(* Logix 5000 project; controller PLC_MCC1300_75F1 vendor 1 type 14 code 166 rev 32.11; software revision 32.04; part 52 of 83 *)
(* tags used below, declared in another part *)
   CONST_rgdDestMask : DINT[32];   // Destination Mask
   CONST_tPlant : UDT_PLANT_CONSTANTS;
   GP_TrackingSearchPlate : GP_TrackingSearchPlate;
   GP_TrackingValidateIndex : GP_TrackingValidateIndex;
   M310_M1_DR_R1 : AXIS_CIP_DRIVE;
   M310_xReqStopPrevConvForPos : BOOL;
   M310Popup : MAC_Popup_ZC[2];
   M310Popup_HMW : MAC_Popup_ZC_HMW[2];
   M310Popup_PlateFreeTimeout : TIMER;
   M310Popup_xDrivePosEnable : BOOL;
   TMP_d : DINT;
   TMP_dDiffPhotocellStartConv0 : DINT;
   TMP_dEndSearch0 : DINT;
   TMP_dEndSearch1 : DINT;
   TMP_dFixedSideOffsetBoth : DINT;
   TMP_dFixedSideOffsetConvoy : DINT;
   TMP_dFixedSideOffsetDW : DINT;
   TMP_dFixedSideOffsetUP : DINT;
   TMP_dHalfConveyorLength : DINT;
   TMP_dHalfPlateLength : DINT;
   TMP_dIndex : DINT;
   TMP_dStartSearch0 : DINT;
   TMP_dStartSearch1 : DINT;
   TMP_xALLForSideLeg : BOOL;
   TMP_xAllLiteToCullet : BOOL;
   TMP_xAtLeastOneForSideLeg : BOOL;
   TMP_xAtLeastOneToCullet : BOOL;
   TMP_xPosHead : BOOL;
   xAlwaysOFF : BOOL;
   xAlwaysON : BOOL;
   xDebugOFF : BOOL;
   Z300_BufferPlate : UDT_LINE_BUFFER_PLATE;
   Z300_Conveyor : UDT_StandConv[29];
   Z300_Conveyor_IN_MOTION : MAC_Conveyor_ZC_IN_MOTION[29];
   Z300_Conveyor_OUT_MOTION : MAC_Conveyor_ZC_OUT_MOTION[29];
   Z300_LineTracking : UDT_LINE_TRACKING;
(* MainProgram, continued *)

ROUTINE M310PopupManagement   (* ladder *)
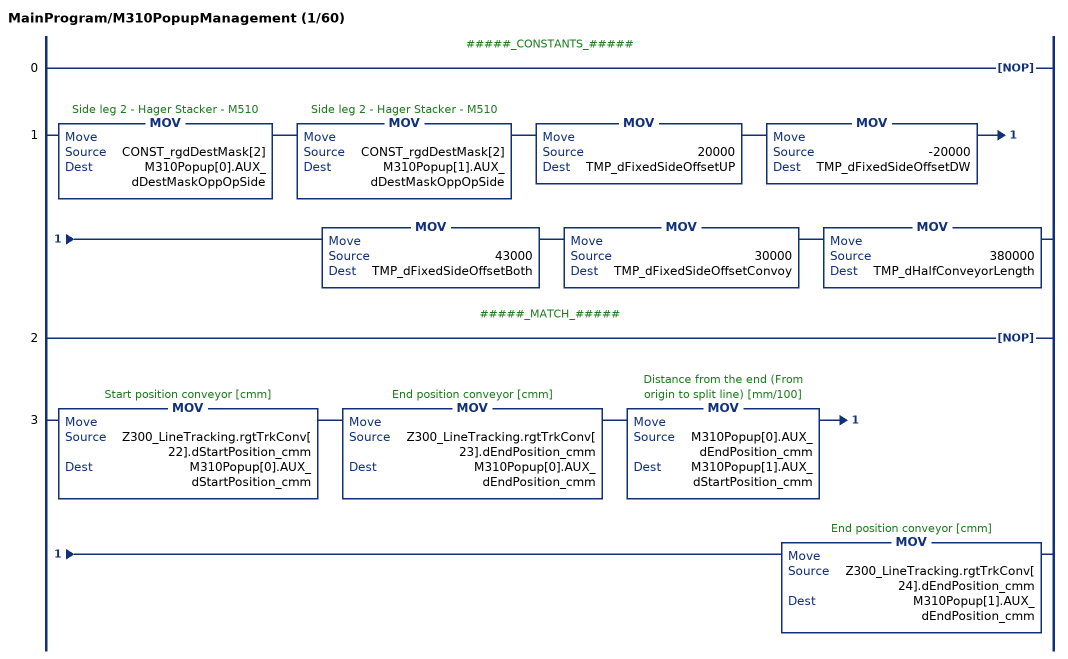
   // #####_CONSTANTS_#####
   0: NOP();
   1: MOV(CONST_rgdDestMask[2],M310Popup[0].AUX_dDestMaskOppOpSide)MOV(CONST_rgdDestMask[2],M310Popup[1].AUX_dDestMaskOppOpSide)MOV(20000,TMP_dFixedSideOffsetUP)MOV(-20000,TMP_dFixedSideOffsetDW)MOV(43000,TMP_dFixedSideOffsetBoth)MOV(30000,TMP_dFixedSideOffsetConvoy)MOV(380000,TMP_dHalfConveyorLength);
   // #####_MATCH_#####
   2: NOP();
   3: MOV(Z300_LineTracking.rgtTrkConv[22].dStartPosition_cmm,M310Popup[0].AUX_dStartPosition_cmm)MOV(Z300_LineTracking.rgtTrkConv[23].dEndPosition_cmm,M310Popup[0].AUX_dEndPosition_cmm)MOV(M310Popup[0].AUX_dEndPosition_cmm,M310Popup[1].AUX_dStartPosition_cmm)MOV(Z300_LineTracking.rgtTrkConv[24].dEndPosition_cmm,M310Popup[1].AUX_dEndPosition_cmm);
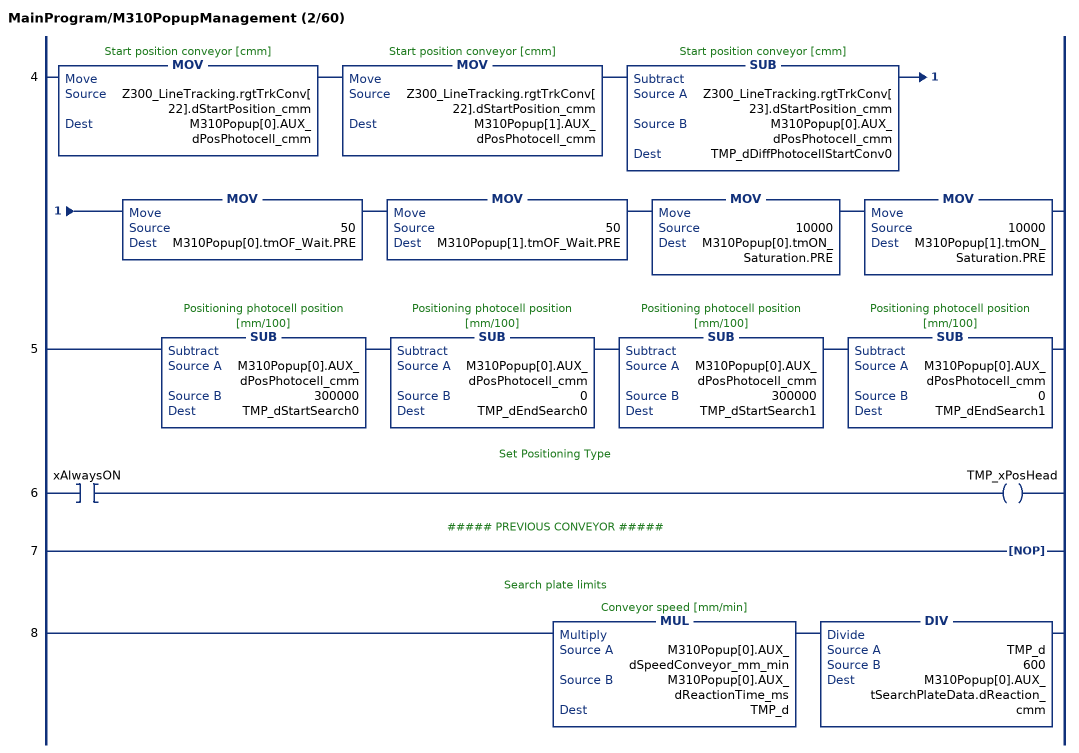
   4: MOV(Z300_LineTracking.rgtTrkConv[22].dStartPosition_cmm,M310Popup[0].AUX_dPosPhotocell_cmm)MOV(Z300_LineTracking.rgtTrkConv[22].dStartPosition_cmm,M310Popup[1].AUX_dPosPhotocell_cmm)SUB(Z300_LineTracking.rgtTrkConv[23].dStartPosition_cmm,M310Popup[0].AUX_dPosPhotocell_cmm,TMP_dDiffPhotocellStartConv0)MOV(50,M310Popup[0].tmOF_Wait.PRE)MOV(50,M310Popup[1].tmOF_Wait.PRE)MOV(10000,M310Popup[0].tmON_Saturation.PRE)MOV(10000,M310Popup[1].tmON_Saturation.PRE);
   5: SUB(M310Popup[0].AUX_dPosPhotocell_cmm,300000,TMP_dStartSearch0)SUB(M310Popup[0].AUX_dPosPhotocell_cmm,0,TMP_dEndSearch0)SUB(M310Popup[0].AUX_dPosPhotocell_cmm,300000,TMP_dStartSearch1)SUB(M310Popup[0].AUX_dPosPhotocell_cmm,0,TMP_dEndSearch1);
   // Set Positioning Type
   6: XIC(xAlwaysON)OTE(TMP_xPosHead);
   // ##### PREVIOUS CONVEYOR #####
   7: NOP();
   // Search plate limits
   8: MUL(M310Popup[0].AUX_dSpeedConveyor_mm_min,M310Popup[0].AUX_dReactionTime_ms,TMP_d)DIV(TMP_d,600,M310Popup[0].AUX_tSearchPlateData.dReaction_cmm);
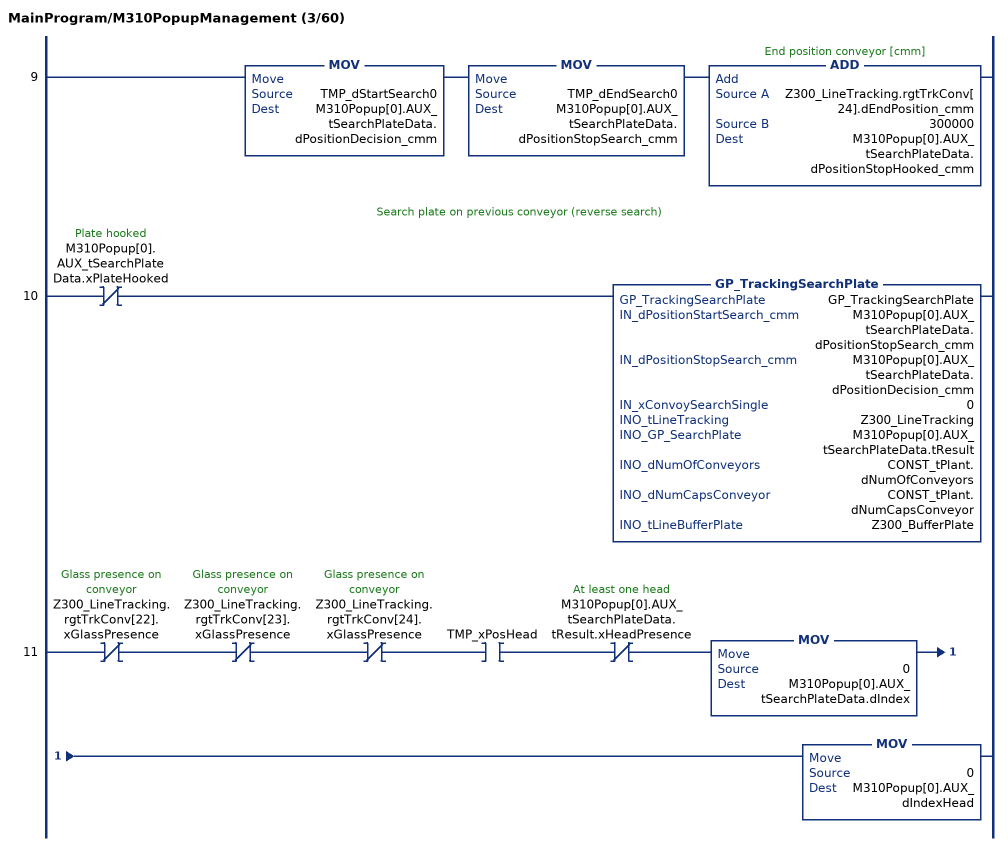
   9: MOV(TMP_dStartSearch0,M310Popup[0].AUX_tSearchPlateData.dPositionDecision_cmm)MOV(TMP_dEndSearch0,M310Popup[0].AUX_tSearchPlateData.dPositionStopSearch_cmm)ADD(Z300_LineTracking.rgtTrkConv[24].dEndPosition_cmm,300000,M310Popup[0].AUX_tSearchPlateData.dPositionStopHooked_cmm);
   // Search plate on previous conveyor (reverse search)
   10: XIO(M310Popup[0].AUX_tSearchPlateData.xPlateHooked)GP_TrackingSearchPlate(GP_TrackingSearchPlate,M310Popup[0].AUX_tSearchPlateData.dPositionStopSearch_cmm,M310Popup[0].AUX_tSearchPlateData.dPositionDecision_cmm,0,Z300_LineTracking,M310Popup[0].AUX_tSearchPlateData.tResult,CONST_tPlant.dNumOfConveyors,CONST_tPlant.dNumCapsConveyor,Z300_BufferPlate);
   11: XIO(Z300_LineTracking.rgtTrkConv[22].xGlassPresence)XIO(Z300_LineTracking.rgtTrkConv[23].xGlassPresence)XIO(Z300_LineTracking.rgtTrkConv[24].xGlassPresence)XIC(TMP_xPosHead)XIO(M310Popup[0].AUX_tSearchPlateData.tResult.xHeadPresence)MOV(0,M310Popup[0].AUX_tSearchPlateData.dIndex)MOV(0,M310Popup[0].AUX_dIndexHead);
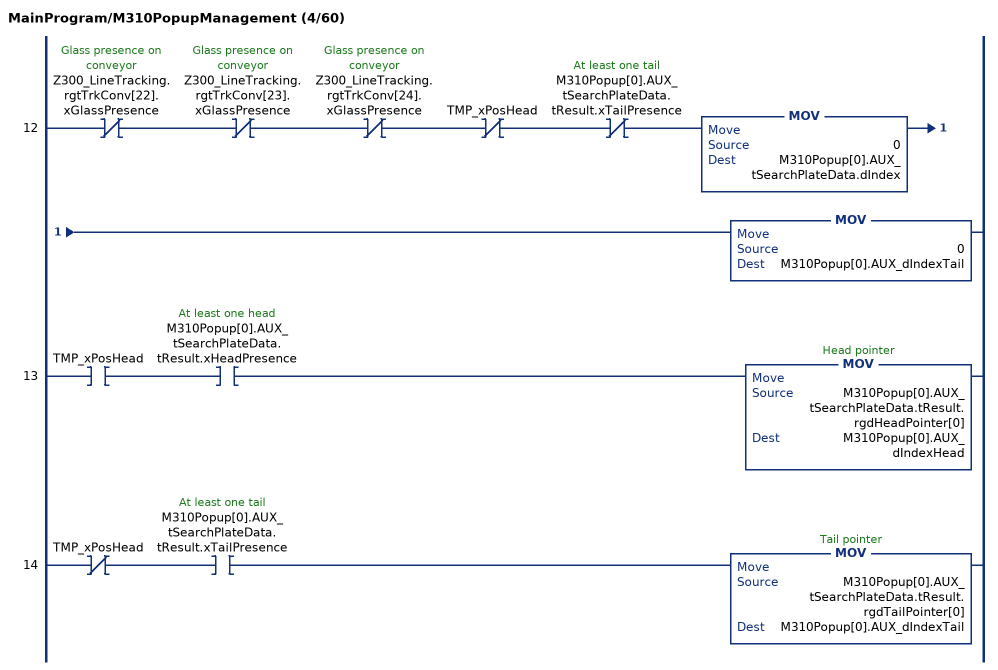
   12: XIO(Z300_LineTracking.rgtTrkConv[22].xGlassPresence)XIO(Z300_LineTracking.rgtTrkConv[23].xGlassPresence)XIO(Z300_LineTracking.rgtTrkConv[24].xGlassPresence)XIO(TMP_xPosHead)XIO(M310Popup[0].AUX_tSearchPlateData.tResult.xTailPresence)MOV(0,M310Popup[0].AUX_tSearchPlateData.dIndex)MOV(0,M310Popup[0].AUX_dIndexTail);
   13: XIC(TMP_xPosHead)XIC(M310Popup[0].AUX_tSearchPlateData.tResult.xHeadPresence)MOV(M310Popup[0].AUX_tSearchPlateData.tResult.rgdHeadPointer[0],M310Popup[0].AUX_dIndexHead);
   14: XIO(TMP_xPosHead)XIC(M310Popup[0].AUX_tSearchPlateData.tResult.xTailPresence)MOV(M310Popup[0].AUX_tSearchPlateData.tResult.rgdTailPointer[0],M310Popup[0].AUX_dIndexTail);
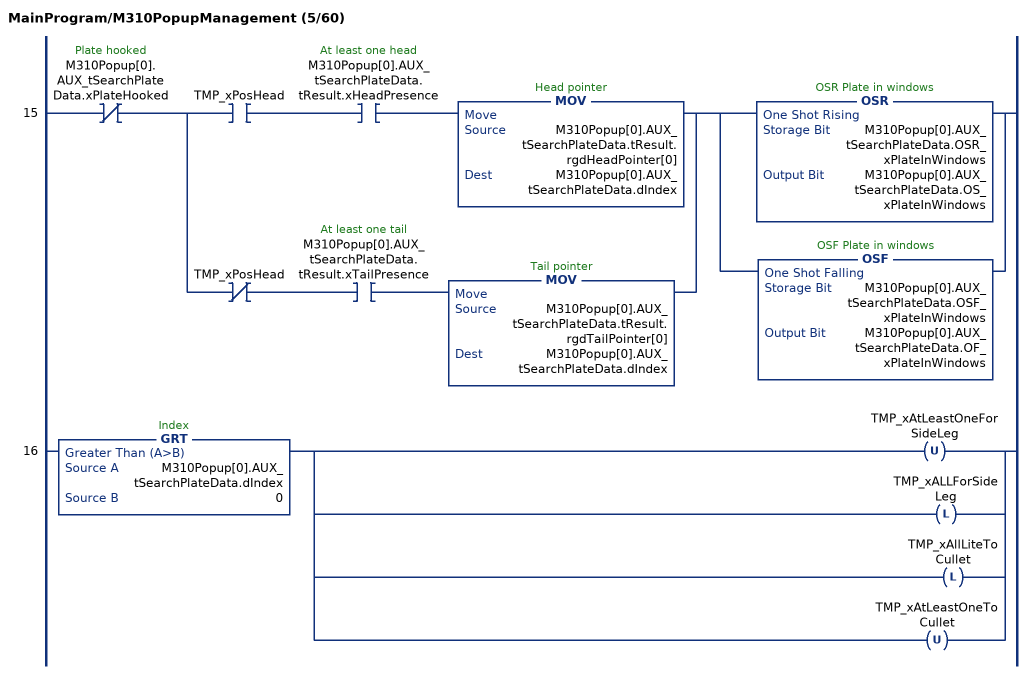
   15: XIO(M310Popup[0].AUX_tSearchPlateData.xPlateHooked)[XIC(TMP_xPosHead) XIC(M310Popup[0].AUX_tSearchPlateData.tResult.xHeadPresence) MOV(M310Popup[0].AUX_tSearchPlateData.tResult.rgdHeadPointer[0],M310Popup[0].AUX_tSearchPlateData.dIndex) ,XIO(TMP_xPosHead) XIC(M310Popup[0].AUX_tSearchPlateData.tResult.xTailPresence) MOV(M310Popup[0].AUX_tSearchPlateData.tResult.rgdTailPointer[0],M310Popup[0].AUX_tSearchPlateData.dIndex) ][OSR(M310Popup[0].AUX_tSearchPlateData.OSR_xPlateInWindows,M310Popup[0].AUX_tSearchPlateData.OS_xPlateInWindows) ,OSF(M310Popup[0].AUX_tSearchPlateData.OSF_xPlateInWindows,M310Popup[0].AUX_tSearchPlateData.OF_xPlateInWindows) ];
   16: GRT(M310Popup[0].AUX_tSearchPlateData.dIndex,0)[OTU(TMP_xAtLeastOneForSideLeg) ,OTL(TMP_xALLForSideLeg) ,OTL(TMP_xAllLiteToCullet) ,OTU(TMP_xAtLeastOneToCullet) ];
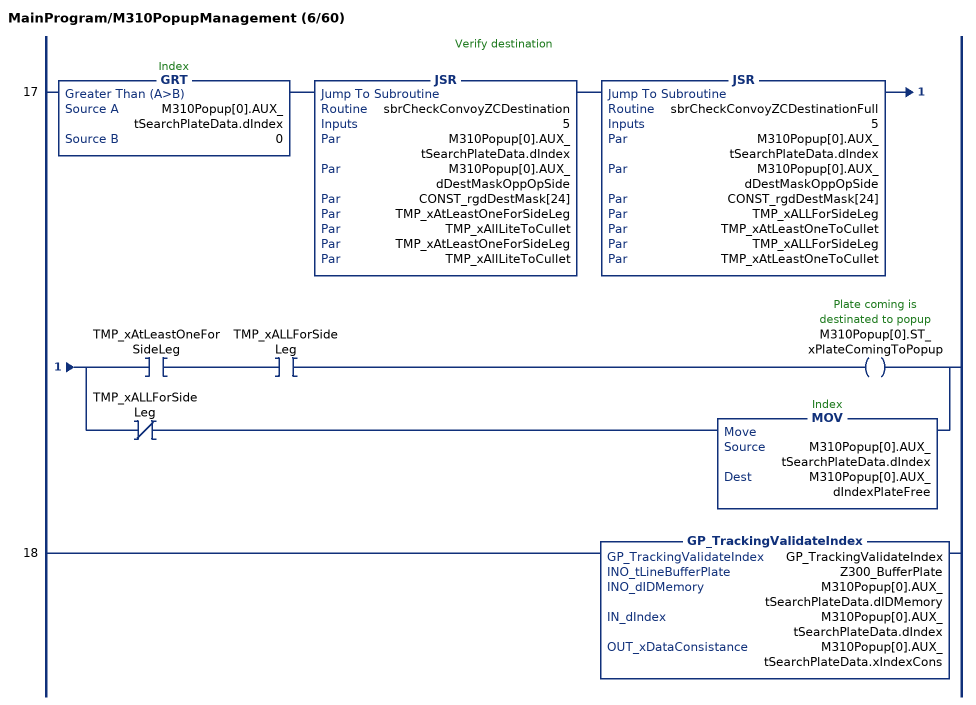
   // Verify destination
   17: GRT(M310Popup[0].AUX_tSearchPlateData.dIndex,0)JSR(sbrCheckConvoyZCDestination,5,M310Popup[0].AUX_tSearchPlateData.dIndex,M310Popup[0].AUX_dDestMaskOppOpSide,CONST_rgdDestMask[24],TMP_xAtLeastOneForSideLeg,TMP_xAllLiteToCullet,TMP_xAtLeastOneForSideLeg,TMP_xAllLiteToCullet)JSR(sbrCheckConvoyZCDestinationFull,5,M310Popup[0].AUX_tSearchPlateData.dIndex,M310Popup[0].AUX_dDestMaskOppOpSide,CONST_rgdDestMask[24],TMP_xALLForSideLeg,TMP_xAtLeastOneToCullet,TMP_xALLForSideLeg,TMP_xAtLeastOneToCullet)[XIC(TMP_xAtLeastOneForSideLeg) XIC(TMP_xALLForSideLeg) OTE(M310Popup[0].ST_xPlateComingToPopup) ,XIO(TMP_xALLForSideLeg) MOV(M310Popup[0].AUX_tSearchPlateData.dIndex,M310Popup[0].AUX_dIndexPlateFree) ];
   18: GP_TrackingValidateIndex(GP_TrackingValidateIndex,Z300_BufferPlate,M310Popup[0].AUX_tSearchPlateData.dIDMemory,M310Popup[0].AUX_tSearchPlateData.dIndex,M310Popup[0].AUX_tSearchPlateData.xIndexCons);
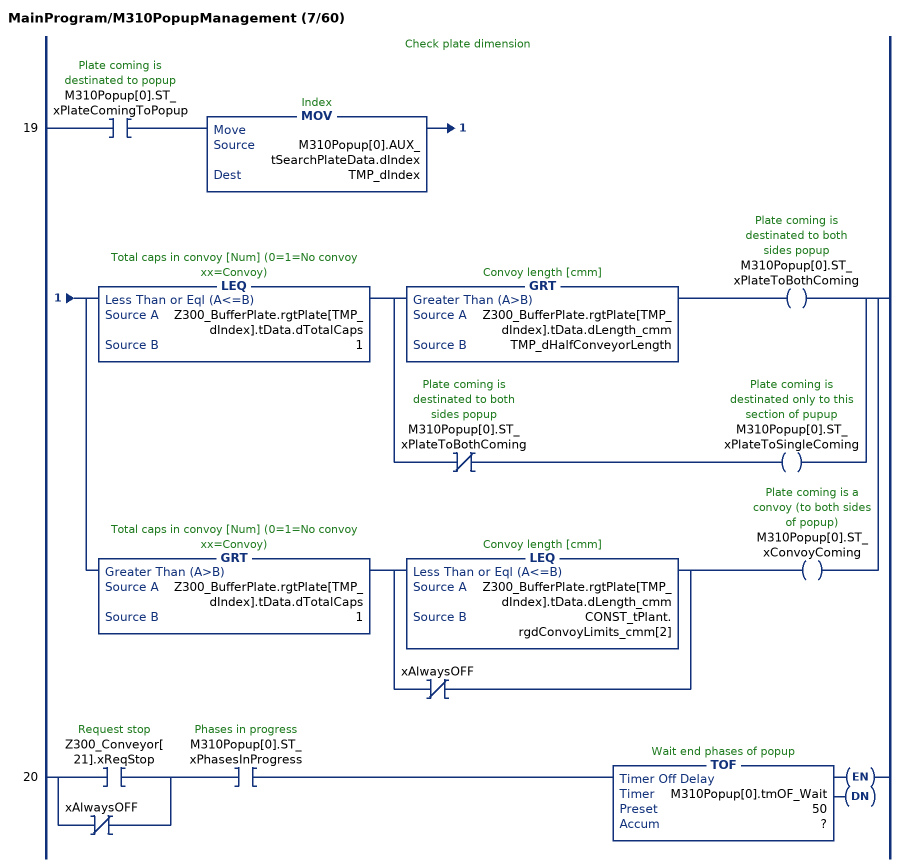
   // Check plate dimension
   19: XIC(M310Popup[0].ST_xPlateComingToPopup)MOV(M310Popup[0].AUX_tSearchPlateData.dIndex,TMP_dIndex)[LEQ(Z300_BufferPlate.rgtPlate[TMP_dIndex].tData.dTotalCaps,1) [GRT(Z300_BufferPlate.rgtPlate[TMP_dIndex].tData.dLength_cmm,TMP_dHalfConveyorLength) OTE(M310Popup[0].ST_xPlateToBothComing) ,XIO(M310Popup[0].ST_xPlateToBothComing) OTE(M310Popup[0].ST_xPlateToSingleComing) ] ,GRT(Z300_BufferPlate.rgtPlate[TMP_dIndex].tData.dTotalCaps,1) [LEQ(Z300_BufferPlate.rgtPlate[TMP_dIndex].tData.dLength_cmm,CONST_tPlant.rgdConvoyLimits_cmm[2]) ,XIO(xAlwaysOFF) ] OTE(M310Popup[0].ST_xConvoyComing) ];
   20: [XIC(Z300_Conveyor[21].xReqStop) ,XIO(xAlwaysOFF) ]XIC(M310Popup[0].ST_xPhasesInProgress)TOF(M310Popup[0].tmOF_Wait,?,?);
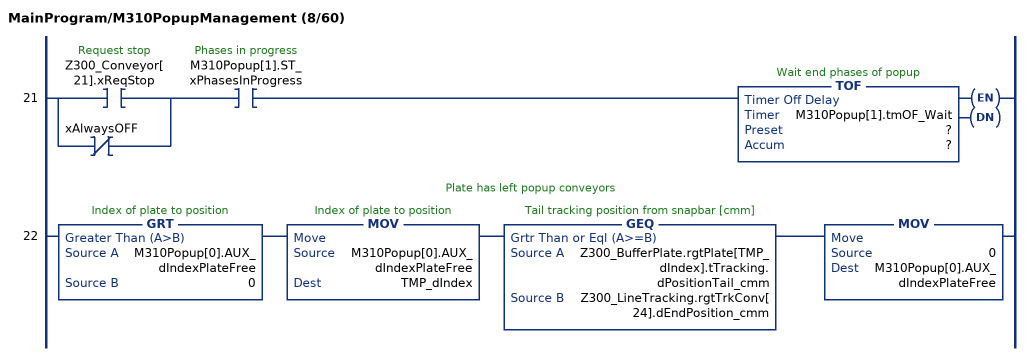
   21: [XIC(Z300_Conveyor[21].xReqStop) ,XIO(xAlwaysOFF) ]XIC(M310Popup[1].ST_xPhasesInProgress)TOF(M310Popup[1].tmOF_Wait,?,?);
   // Plate has left popup conveyors
   22: GRT(M310Popup[0].AUX_dIndexPlateFree,0)MOV(M310Popup[0].AUX_dIndexPlateFree,TMP_dIndex)GEQ(Z300_BufferPlate.rgtPlate[TMP_dIndex].tTracking.dPositionTail_cmm,Z300_LineTracking.rgtTrkConv[24].dEndPosition_cmm)MOV(0,M310Popup[0].AUX_dIndexPlateFree);
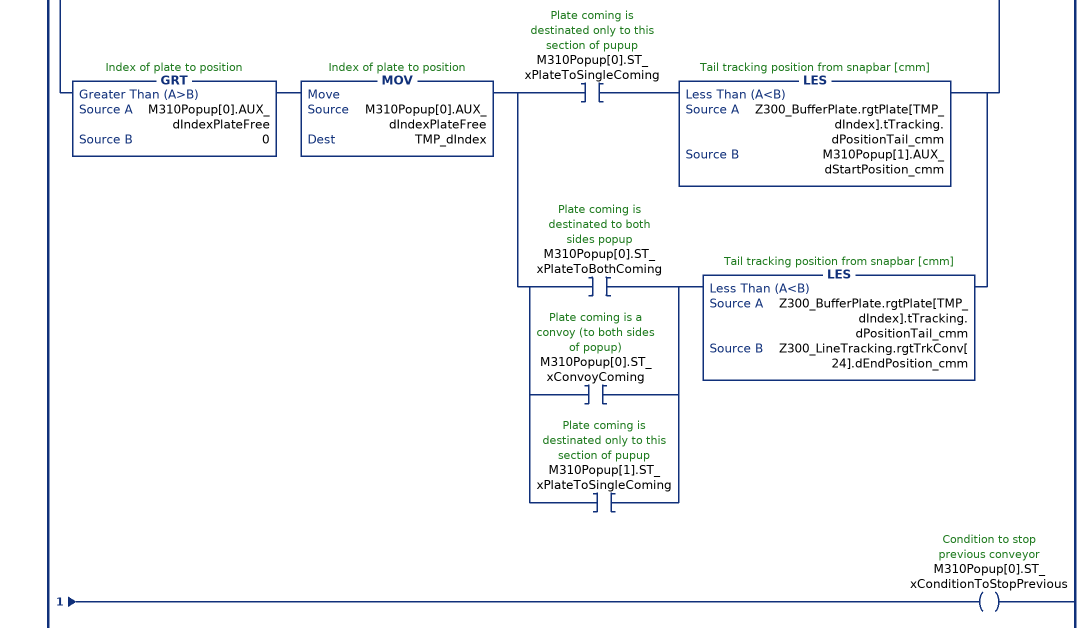
   // Stop previuos conveyor if no condition on pop-up conveyor
   23: [[XIC(M310Popup[0].ST_xPlateToSingleComing) [XIO(M310Popup[0].ST_xInitialConditionForRise) ,XIC(M310Popup[0].ST_xPlatePresentOnPopup) ,XIC(M310Popup[0].ST_xPlatePresence) ,XIC(Z300_LineTracking.rgtTrkConv[22].xGlassPresence) ,XIC(Z300_LineTracking.rgtTrkConv[23].xGlassPresence) ,EQU(M310Popup[0].AUX_dIndexPositioning,0) [XIC(M310Popup[0].ST_xPlateUnderPopup) ,XIC(M310Popup[1].ST_xPlateUnderPopup) ] ] ,XIC(M310Popup[0].ST_xPlateToSingleComing) [XIO(M310Popup[1].ST_xInitialConditionForRise) ,XIC(M310Popup[1].ST_xPlatePresentOnPopup) ,XIC(M310Popup[1].ST_xPlatePresence) ,XIC(Z300_LineTracking.rgtTrkConv[22].xGlassPresence) ,XIC(Z300_LineTracking.rgtTrkConv[23].xGlassPresence) ,XIC(Z300_LineTracking.rgtTrkConv[24].xGlassPresence) ,EQU(M310Popup[0].AUX_dIndexPositioning,0) [XIC(M310Popup[0].ST_xPlateUnderPopup) ,XIC(M310Popup[1].ST_xPlateUnderPopup) ] ] ,[XIC(M310Popup[0].ST_xPlateToBothComing) ,XIC(M310Popup[0].ST_xConvoyComing) ] [XIO(M310Popup[1].ST_xInitialConditionForRise) ,XIC(M310Popup[1].ST_xPlatePresentOnPopup) ,XIC(M310Popup[1].ST_xPlatePresence) ,XIC(Z300_LineTracking.rgtTrkConv[22].xGlassPresence) ,XIC(Z300_LineTracking.rgtTrkConv[23].xGlassPresence) ,XIC(Z300_LineTracking.rgtTrkConv[24].xGlassPresence) ,EQU(M310Popup[0].AUX_dIndexPositioning,0) XIC(M310Popup[1].ST_xPlateUnderPopup) ,XIO(M310Popup[0].ST_xInitialConditionForRise) ,XIC(M310Popup[0].ST_xPlatePresentOnPopup) ,XIC(M310Popup[0].ST_xPlatePresence) ,EQU(M310Popup[0].AUX_dIndexPositioning,0) XIC(M310Popup[0].ST_xPlateUnderPopup) ] ] ,XIO(M310Popup[0].INPUT_xPopupHigh) XIO(M310Popup[0].INPUT_xPopupLow) ,XIO(M310Popup[1].INPUT_xPopupHigh) XIO(M310Popup[1].INPUT_xPopupLow) ,XIC(M310_xReqStopPrevConvForPos) ,XIC(Z300_Conveyor[22].xReqExtStopLoadNewPlate) ,[XIC(M310Popup[0].ST_xPlateInPositionToRise) ,XIC(M310Popup[1].ST_xPlateInPositionToRise) ] ,XIC(Z300_Conveyor[22].ST_xCleaningEnabled) XIO(Z300_Conveyor[21].ST_xCleaningEnabled) ,XIC(M310Popup[0].ST_xPrevConvFreeAfterPos) ,XIC(M310Popup[1].ST_xPrevConvFreeAfterPos) ,[XIO(M310Popup[0].INPUT_xPopupHigh) ,XIO(M310Popup[1].INPUT_xPopupHigh) ] ,GRT(M310Popup[0].AUX_dIndexPositioning,0) [GRT(M310Popup[0].AUX_tSearchPlateData.dIndex,0) NEQ(M310Popup[0].AUX_tSearchPlateData.dIndex,M310Popup[0].AUX_dIndexPositioning) ,GRT(M310Popup[0].AUX_dIndexPlatePositioned,0) NEQ(M310Popup[0].AUX_dIndexPlatePositioned,M310Popup[0].AUX_dIndexPositioning) ] ,GRT(M310Popup[0].AUX_dIndexPlateFree,0) MOV(M310Popup[0].AUX_dIndexPlateFree,TMP_dIndex) [XIC(M310Popup[0].ST_xPlateToSingleComing) LES(Z300_BufferPlate.rgtPlate[TMP_dIndex].tTracking.dPositionTail_cmm,M310Popup[1].AUX_dStartPosition_cmm) ,[XIC(M310Popup[0].ST_xPlateToBothComing) ,XIC(M310Popup[0].ST_xConvoyComing) ,XIC(M310Popup[1].ST_xPlateToSingleComing) ] LES(Z300_BufferPlate.rgtPlate[TMP_dIndex].tTracking.dPositionTail_cmm,Z300_LineTracking.rgtTrkConv[24].dEndPosition_cmm) ] ]OTE(M310Popup[0].ST_xConditionToStopPrevious);
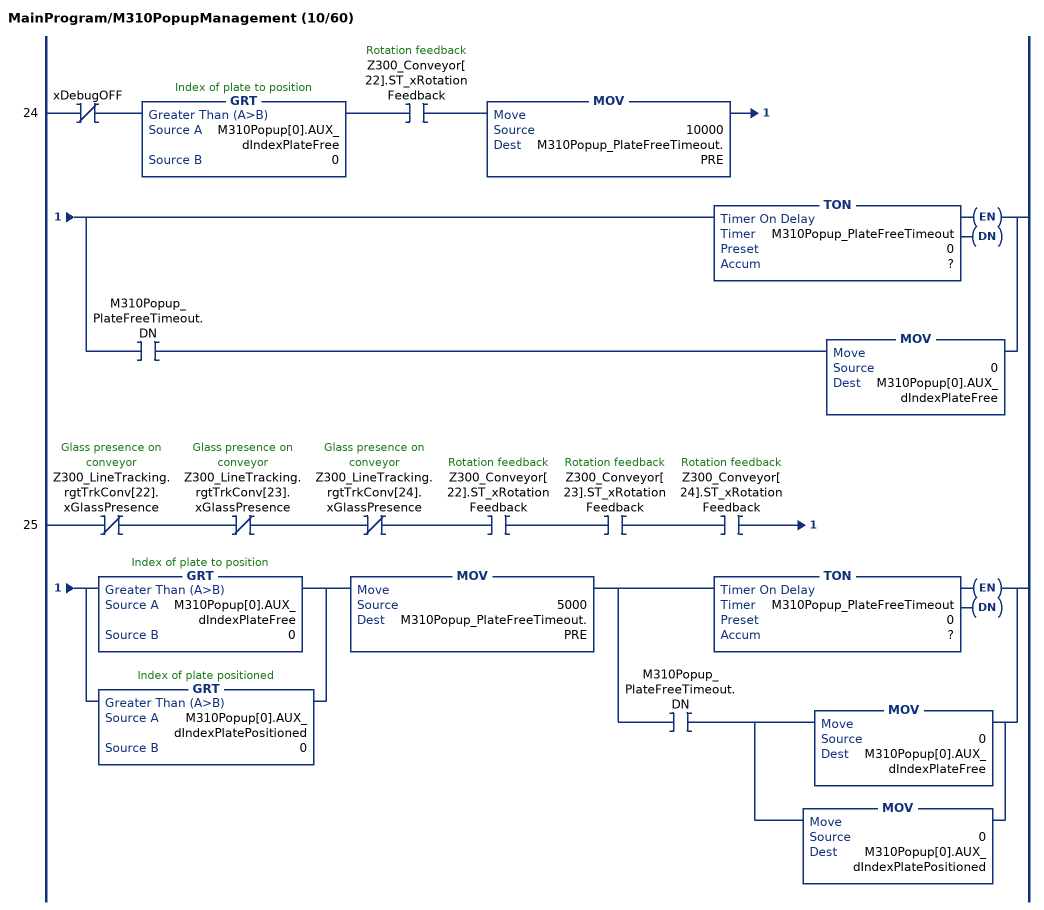
   24: XIO(xDebugOFF)GRT(M310Popup[0].AUX_dIndexPlateFree,0)XIC(Z300_Conveyor[22].ST_xRotationFeedback)MOV(10000,M310Popup_PlateFreeTimeout.PRE)[TON(M310Popup_PlateFreeTimeout,?,?) ,XIC(M310Popup_PlateFreeTimeout.DN) MOV(0,M310Popup[0].AUX_dIndexPlateFree) ];
   25: XIO(Z300_LineTracking.rgtTrkConv[22].xGlassPresence)XIO(Z300_LineTracking.rgtTrkConv[23].xGlassPresence)XIO(Z300_LineTracking.rgtTrkConv[24].xGlassPresence)XIC(Z300_Conveyor[22].ST_xRotationFeedback)XIC(Z300_Conveyor[23].ST_xRotationFeedback)XIC(Z300_Conveyor[24].ST_xRotationFeedback)[GRT(M310Popup[0].AUX_dIndexPlateFree,0) ,GRT(M310Popup[0].AUX_dIndexPlatePositioned,0) ]MOV(5000,M310Popup_PlateFreeTimeout.PRE)[TON(M310Popup_PlateFreeTimeout,?,?) ,XIC(M310Popup_PlateFreeTimeout.DN) [MOV(0,M310Popup[0].AUX_dIndexPlateFree) ,MOV(0,M310Popup[0].AUX_dIndexPlatePositioned) ] ];
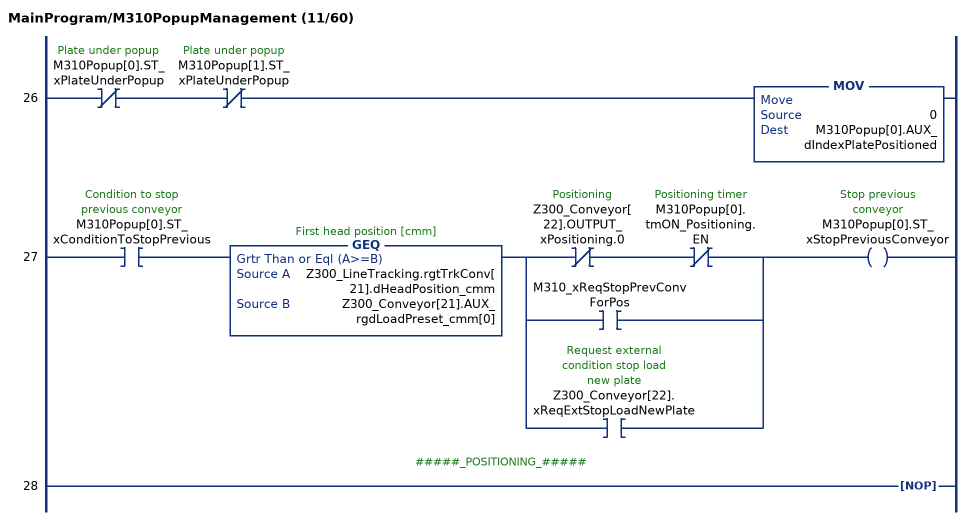
   26: XIO(M310Popup[0].ST_xPlateUnderPopup)XIO(M310Popup[1].ST_xPlateUnderPopup)MOV(0,M310Popup[0].AUX_dIndexPlatePositioned);
   27: XIC(M310Popup[0].ST_xConditionToStopPrevious)GEQ(Z300_LineTracking.rgtTrkConv[21].dHeadPosition_cmm,Z300_Conveyor[21].AUX_rgdLoadPreset_cmm[0])[XIO(Z300_Conveyor[22].OUTPUT_xPositioning.0) XIO(M310Popup[0].tmON_Positioning.EN) ,[XIC(M310_xReqStopPrevConvForPos) ,XIC(Z300_Conveyor[22].xReqExtStopLoadNewPlate) ] ]OTE(M310Popup[0].ST_xStopPreviousConveyor);
   // #####_POSITIONING_#####
   28: NOP();
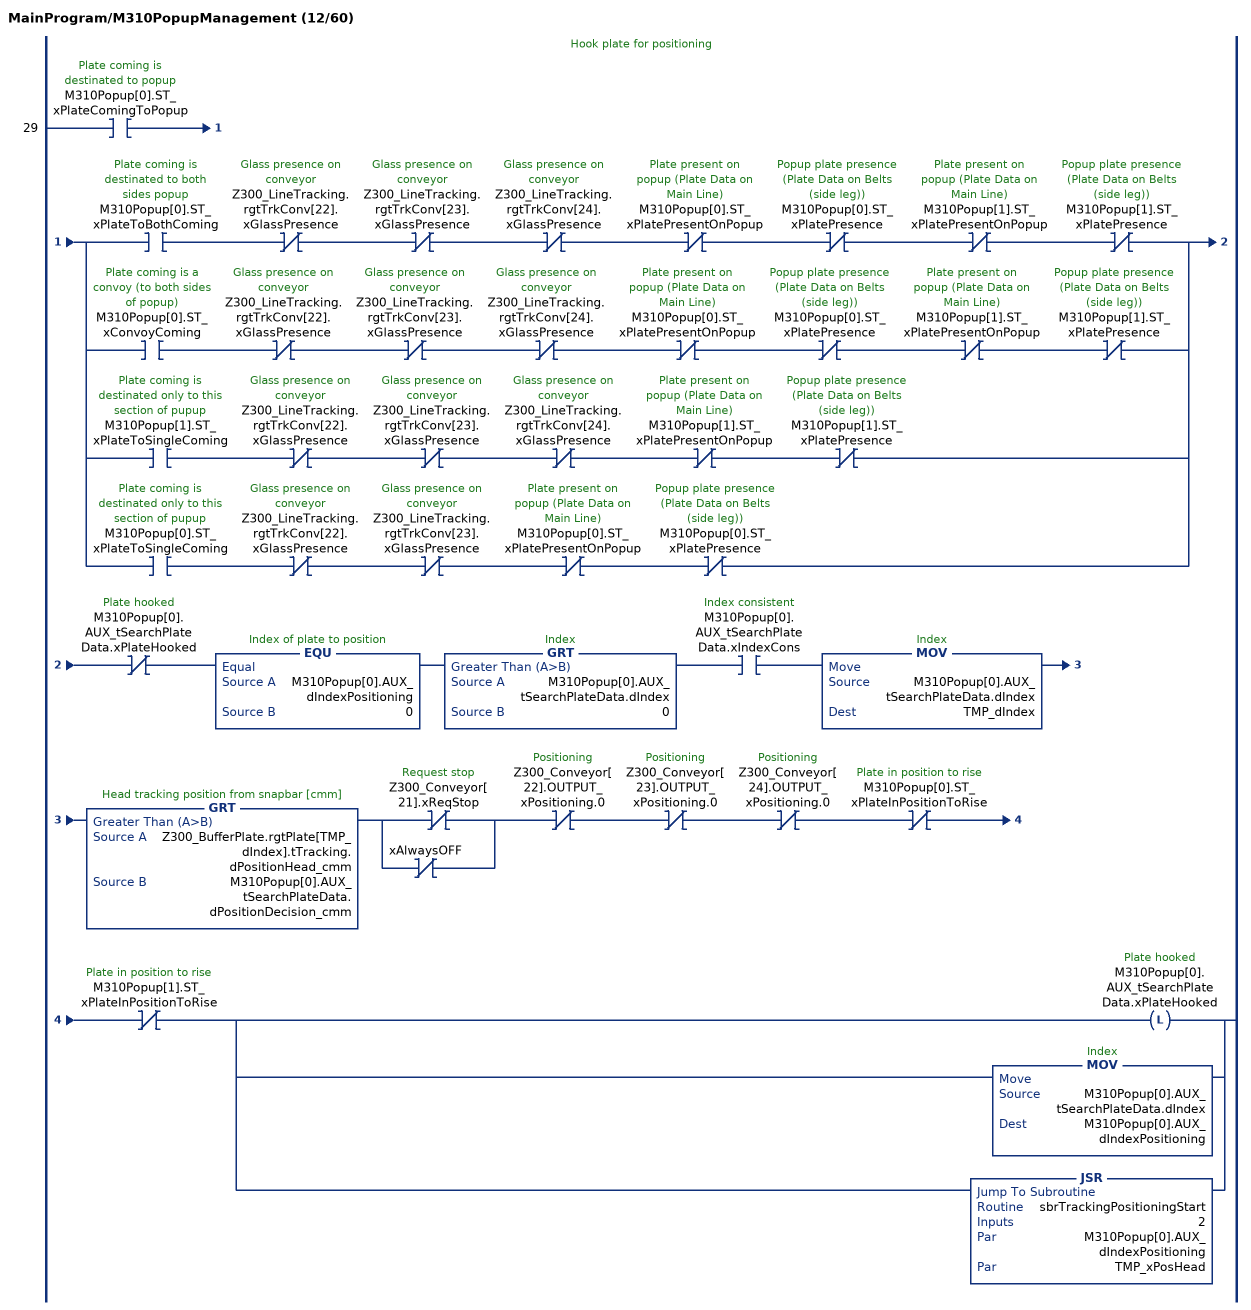
   // Hook plate for positioning
   29: XIC(M310Popup[0].ST_xPlateComingToPopup)[XIC(M310Popup[0].ST_xPlateToBothComing) XIO(Z300_LineTracking.rgtTrkConv[22].xGlassPresence) XIO(Z300_LineTracking.rgtTrkConv[23].xGlassPresence) XIO(Z300_LineTracking.rgtTrkConv[24].xGlassPresence) XIO(M310Popup[0].ST_xPlatePresentOnPopup) XIO(M310Popup[0].ST_xPlatePresence) XIO(M310Popup[1].ST_xPlatePresentOnPopup) XIO(M310Popup[1].ST_xPlatePresence) ,XIC(M310Popup[0].ST_xConvoyComing) XIO(Z300_LineTracking.rgtTrkConv[22].xGlassPresence) XIO(Z300_LineTracking.rgtTrkConv[23].xGlassPresence) XIO(Z300_LineTracking.rgtTrkConv[24].xGlassPresence) XIO(M310Popup[0].ST_xPlatePresentOnPopup) XIO(M310Popup[0].ST_xPlatePresence) XIO(M310Popup[1].ST_xPlatePresentOnPopup) XIO(M310Popup[1].ST_xPlatePresence) ,XIC(M310Popup[1].ST_xPlateToSingleComing) XIO(Z300_LineTracking.rgtTrkConv[22].xGlassPresence) XIO(Z300_LineTracking.rgtTrkConv[23].xGlassPresence) XIO(Z300_LineTracking.rgtTrkConv[24].xGlassPresence) XIO(M310Popup[1].ST_xPlatePresentOnPopup) XIO(M310Popup[1].ST_xPlatePresence) ,XIC(M310Popup[0].ST_xPlateToSingleComing) XIO(Z300_LineTracking.rgtTrkConv[22].xGlassPresence) XIO(Z300_LineTracking.rgtTrkConv[23].xGlassPresence) XIO(M310Popup[0].ST_xPlatePresentOnPopup) XIO(M310Popup[0].ST_xPlatePresence) ]XIO(M310Popup[0].AUX_tSearchPlateData.xPlateHooked)EQU(M310Popup[0].AUX_dIndexPositioning,0)GRT(M310Popup[0].AUX_tSearchPlateData.dIndex,0)XIC(M310Popup[0].AUX_tSearchPlateData.xIndexCons)MOV(M310Popup[0].AUX_tSearchPlateData.dIndex,TMP_dIndex)GRT(Z300_BufferPlate.rgtPlate[TMP_dIndex].tTracking.dPositionHead_cmm,M310Popup[0].AUX_tSearchPlateData.dPositionDecision_cmm)[XIO(Z300_Conveyor[21].xReqStop) ,XIO(xAlwaysOFF) ]XIO(Z300_Conveyor[22].OUTPUT_xPositioning.0)XIO(Z300_Conveyor[23].OUTPUT_xPositioning.0)XIO(Z300_Conveyor[24].OUTPUT_xPositioning.0)XIO(M310Popup[0].ST_xPlateInPositionToRise)XIO(M310Popup[1].ST_xPlateInPositionToRise)[OTL(M310Popup[0].AUX_tSearchPlateData.xPlateHooked) ,MOV(M310Popup[0].AUX_tSearchPlateData.dIndex,M310Popup[0].AUX_dIndexPositioning) ,JSR(sbrTrackingPositioningStart,2,M310Popup[0].AUX_dIndexPositioning,TMP_xPosHead) ];
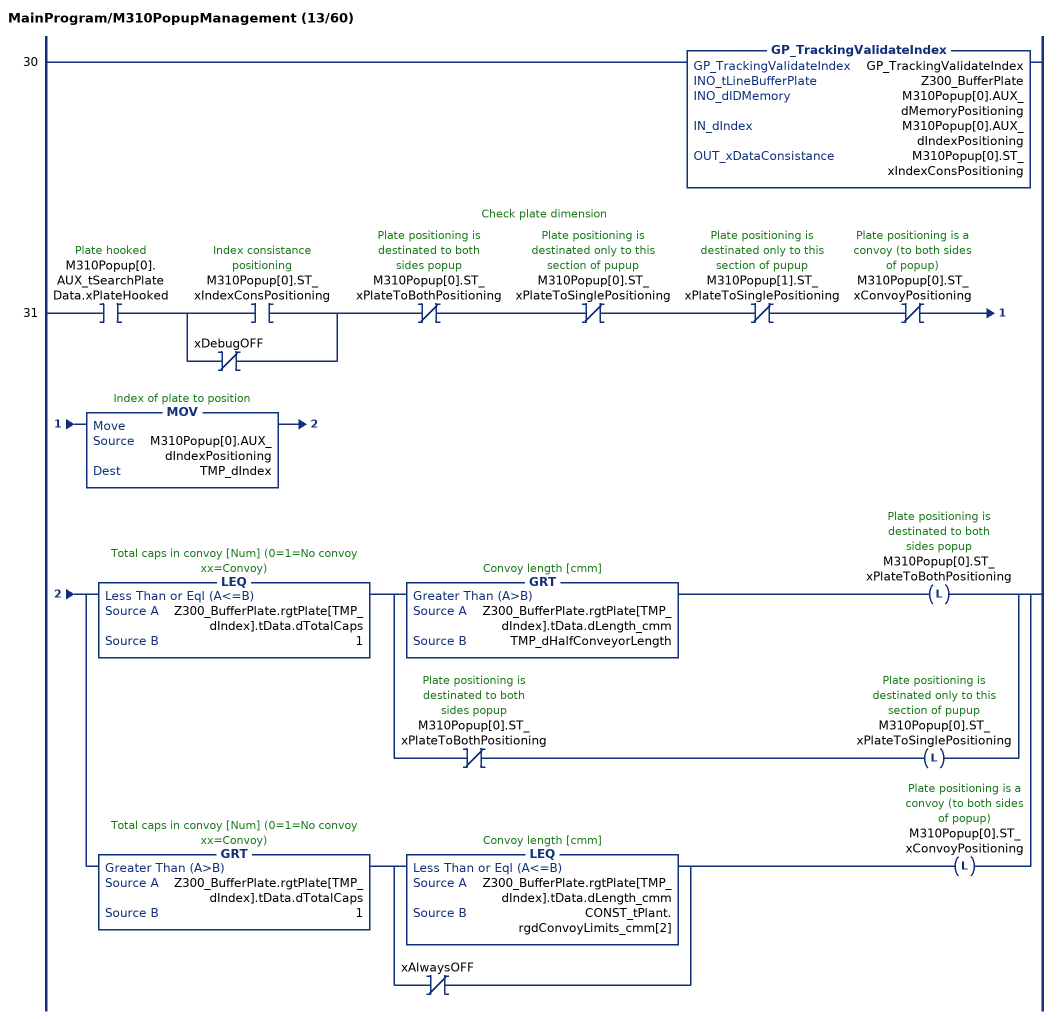
   30: GP_TrackingValidateIndex(GP_TrackingValidateIndex,Z300_BufferPlate,M310Popup[0].AUX_dMemoryPositioning,M310Popup[0].AUX_dIndexPositioning,M310Popup[0].ST_xIndexConsPositioning);
   // Check plate dimension
   31: XIC(M310Popup[0].AUX_tSearchPlateData.xPlateHooked)[XIC(M310Popup[0].ST_xIndexConsPositioning) ,XIO(xDebugOFF) ]XIO(M310Popup[0].ST_xPlateToBothPositioning)XIO(M310Popup[0].ST_xPlateToSinglePositioning)XIO(M310Popup[1].ST_xPlateToSinglePositioning)XIO(M310Popup[0].ST_xConvoyPositioning)MOV(M310Popup[0].AUX_dIndexPositioning,TMP_dIndex)[LEQ(Z300_BufferPlate.rgtPlate[TMP_dIndex].tData.dTotalCaps,1) [GRT(Z300_BufferPlate.rgtPlate[TMP_dIndex].tData.dLength_cmm,TMP_dHalfConveyorLength) OTL(M310Popup[0].ST_xPlateToBothPositioning) ,XIO(M310Popup[0].ST_xPlateToBothPositioning) OTL(M310Popup[0].ST_xPlateToSinglePositioning) ] ,GRT(Z300_BufferPlate.rgtPlate[TMP_dIndex].tData.dTotalCaps,1) [LEQ(Z300_BufferPlate.rgtPlate[TMP_dIndex].tData.dLength_cmm,CONST_tPlant.rgdConvoyLimits_cmm[2]) ,XIO(xAlwaysOFF) ] OTL(M310Popup[0].ST_xConvoyPositioning) ];